
screen "3161_ParetoAlarmData" 1280x715, template "3xxx_Alarms&Events"
   Rectangle "recBaseScreenLocked" at 0,0 size 1280x708
      Visibility <- "bo_System_BaseScreenLocked"
   TextField "Text_SortBy" at 33,29 size 102x31; Text 'Sort By:'
   SymbolicIOField "List_ParetoSort" at 135,28 size 244x33; TextOn '1'; TextOff '0'; TextList "Pareto_Sort"
      ProcessValue <- "ParetoData_Sort"
   TextField "Title_Alarm" at 1,84 size 50x21; Text 'Alarm'
   TextField "Title_ID" at 63,84 size 24x21; Text 'ID'
   TextField "Title_Message" at 286,84 size 71x21; Text 'Meldung / Message'
   TextField "Title_TimesOccurred" at 516,67 size 76x38; Text 'Anzahl Time Occurred'
   TextField "Title_TotalDowntime" at 584,67 size 102x38; Text 'Unproduktiv Total Downtime'
   TextField "Title_MTTR" at 682,84 size 49x21; Text 'MTTR'
   TextField "Title_%" at 761,84 size 23x21; Text '%'
   TextField "Text_TotalUptime" at 842,192 size 119x40; Text 'Produktiv: [min] Total Uptime: [min]'
   TextField "Text_TotalDowntime" at 818,250 size 143x40; Text 'Unproduktiv: [min] Total Downtime: [min]'
   TextField "Text_PercentUptime" at 821,316 size 140x22; Text 'Produktiv in %: / Percent Uptime:'
   TextField "Text_TotalStops" at 855,374 size 106x22; Text 'Stopps: / Total Stops:'
   TextField "Text_MTTR" at 903,422 size 58x40; Text 'MTTR: [min]'
   TextField "Text_MTBF" at 904,480 size 57x40; Text 'MTBF: [min]'
   Button "Reset_Button" at 833,539 size 254x32; TextOff 'RESET'
      on Press: function_b14e0dd5("ParetoData_Reset", 0)
   IOField "TotalUptime" at 967,197 size 120x30; FormatPattern 9999.99
      ProcessValue <- "ParetoData_totalUptime"
   IOField "TotalDowntime" at 967,255 size 120x30; FormatPattern 9999.99
      ProcessValue <- "ParetoData_totalDowntime"
   IOField "PercentUptime" at 967,312 size 120x30; FormatPattern 999.9
      ProcessValue <- "ParetoData_percentUptime"
   IOField "TotalStops" at 967,370 size 120x30; FormatPattern 999
      ProcessValue <- "ParetoData_totalStops"
   IOField "MTTR" at 967,427 size 120x30; FormatPattern 9999.99
      ProcessValue <- "ParetoData_MTTR"
   IOField "MTBF" at 967,485 size 120x30; FormatPattern 9999.99
      ProcessValue <- "ParetoData_MTBF"
   TextField "Title_Alarm_1" at 14,118 size 29x31; Text '1:'
   TextField "Title_Alarm_2" at 14,166 size 29x31; Text '2:'
   TextField "Title_Alarm_3" at 14,214 size 29x31; Text '3:'
   TextField "Title_Alarm_4" at 14,262 size 29x31; Text '4:'
   TextField "Title_Alarm_5" at 14,310 size 29x31; Text '5:'
   TextField "Title_Alarm_6" at 14,358 size 29x31; Text '6:'
   TextField "Title_Alarm_7" at 14,406 size 29x31; Text '7:'
   TextField "Title_Alarm_8" at 14,454 size 29x31; Text '8:'
   TextField "Title_Alarm_9" at 14,502 size 29x31; Text '9:'
   TextField "Title_Alarm_10" at 6,550 size 44x31; Text '10:'
   TextField "Text_TotalTimeSinceReset" at 850,126 size 111x58; Text 'Zeit seit Rücksetzen: [min] Total Time Since Reset: [min]'
   IOField "TotalTimeSinceReset" at 967,140 size 120x30; FormatPattern 9999.99
      ProcessValue <- "ParetoData_totalTimeSinceReset"
   ScreenModuleView "ParetoFacePlate_1" at 49,115 size 760x38; ScreenModuleType ""
      Guid_{11997190-103935} <- "ParetoData_alarmOccurrence[1]"
   ScreenModuleView "ParetoFacePlate_2" at 49,163 size 760x38; ScreenModuleType ""
      Guid_{11997190-103935} <- "ParetoData_alarmOccurrence[2]"
   ScreenModuleView "ParetoFacePlate_3" at 49,211 size 760x38; ScreenModuleType ""
      Guid_{11997190-103935} <- "ParetoData_alarmOccurrence[3]"
   ScreenModuleView "ParetoFacePlate_4" at 49,259 size 760x38; ScreenModuleType ""
      Guid_{11997190-103935} <- "ParetoData_alarmOccurrence[4]"
   ScreenModuleView "ParetoFacePlate_5" at 49,307 size 760x38; ScreenModuleType ""
      Guid_{11997190-103935} <- "ParetoData_alarmOccurrence[5]"
   ScreenModuleView "ParetoFacePlate_6" at 49,355 size 760x38; ScreenModuleType ""
      Guid_{11997190-103935} <- "ParetoData_alarmOccurrence[6]"
   ScreenModuleView "ParetoFacePlate_7" at 49,403 size 760x38; ScreenModuleType ""
      Guid_{11997190-103935} <- "ParetoData_alarmOccurrence[7]"
   ScreenModuleView "ParetoFacePlate_8" at 49,451 size 760x38; ScreenModuleType ""
      Guid_{11997190-103935} <- "ParetoData_alarmOccurrence[8]"
   ScreenModuleView "ParetoFacePlate_9" at 49,499 size 760x38; ScreenModuleType ""
      Guid_{11997190-103935} <- "ParetoData_alarmOccurrence[9]"
   ScreenModuleView "ParetoFacePlate_10" at 49,547 size 760x38; ScreenModuleType ""
      Guid_{11997190-103935} <- "ParetoData_alarmOccurrence[10]"

screen "7001_RecipeControl" 1280x715, template "7xxx_Formats"
   Button "btn_Save" at 937,17 size 156x71; TextOff 'Save Current Recipe Datensatz Speichern Salvar'
      on Release: ResetBit("CPG_Recipe_Management.HMI_Command.Save.saveCmd")
      on Press: SetBit("CPG_Recipe_Management.HMI_Command.Save.saveCmd")
   Button "btn_Save_1" at 25,29 size 111x48; TextOff 'Reset All Times Rücksetzen Salvar'
      on Release: ResetBit("CPG_Recipe_Management.HMI_Command.resetAllTimes")
      on Press: SetBit("CPG_Recipe_Management.HMI_Command.resetAllTimes")
   Button "btn_Delete" at 444,538 size 150x45; TextOff 'Change Recipe Datensatz Ändern'
      on Release: ResetBit("CPG_Recipe_Management.HMI_Command.Change.changeCmd")
      on Press: SetBit("CPG_Recipe_Management.HMI_Command.Change.changeCmd")
   Button "btn_Rename" at 607,538 size 150x45; TextOff 'Save Recipe As Datensatz Speichern unter Rebautizar:'
      on Release: ResetBit("CPG_Recipe_Management.HMI_Command.Save.saveAsCmd")
      on Press: SetBit("CPG_Recipe_Management.HMI_Command.Save.saveAsCmd")
   Button "btn_WriteToPLC" at 771,538 size 150x45; TextOff 'Copy Recipe Datensatz Kopieren Write to PLC'
      on Release: ResetBit("CPG_Recipe_Management.HMI_Command.Copy.copyCmd")
      on Press: SetBit("CPG_Recipe_Management.HMI_Command.Copy.copyCmd")
   Button "btn_ReadFromPLC" at 935,538 size 150x45; TextOff 'Delete Recipe Datensatz Löschen Leer desde PLC'
      on Release: ResetBit("CPG_Recipe_Management.HMI_Command.Delete.deleteCmd")
      on Press: SetBit("CPG_Recipe_Management.HMI_Command.Delete.deleteCmd")
   Button "rec_BaseScreenLocked" at 0,0 size 1280x715; TextOff 'Text'
      Visibility <- "bo_System_BaseScreenLocked"
   IOField "I/O field_2" at 345,38 size 38x29; FormatPattern 999
      ProcessValue <- "CurrentRecipeID"
   TextField "Text field_5" at 166,39 size 157x27; Text 'Current Recipe: / Aktueller Datensatz:'
   IOField "I/O field_19" at 171,91 size 189x29; FormatPattern ????????????????????
      ProcessValue <- "CurrentRecipeName"
   TextField "Text field_26" at 8,84 size 156x48; Text 'Tap to Rename Current Recipe: Aktuellen Datensatz Umbenennen:'
   Button "Button_3" at 13,559 size 78x45; TextOff 'Text'; PictureOff "Up_Arrow"
      on Release: function_b9b71300("CPG_Recipe_Management.currentPages[4]", 1)
   Button "Button_4" at 117,559 size 78x45; TextOff 'Text'; PictureOff "Down_Arrow"
      on Release: function_dd21b452("CPG_Recipe_Management.currentPages[4]", 1)
   IOField "I/O field_30" at 293,571 size 35x21; FormatPattern 999
      ProcessValue <- "CPG_Recipe_Management.currentPages[4]"
   TextField "Text field_46" at 225,569 size 60x25; Text 'Page # / Seite #'
   TextField "Text field_47" at 337,569 size 32x25; Text 'of / von'
   IOField "I/O field_45" at 385,572 size 27x19; FormatPattern 999
      ProcessValue <- "CPG_Recipe_Management.maxPages[4]"
   Rectangle "Rectangle_7" at 438,24 size 224x56
      Visibility <- "RecipeChangeDisabled"
   TextField "Text field_45" at 455,28 size 190x48; Text 'Recipe changes disabled due to machine state Änderungen gesperrt wegen Maschinenzustand'
      Visibility <- "RecipeChangeDisabled"
   Rectangle "Rectangle_2" at 668,24 size 261x56
      Visibility <- "RecipeSetpointDiff"
   TextField "Text field_27" at 674,28 size 249x48; Text 'Warning: At least one value differs from the saved setpoints! Mindestens ein Wert entspricht nicht den Speicherwerten!'
      Visibility <- "RecipeSetpointDiff"
   Group "Group" at 5,531 size 421x27
   Group "Group_1" at 5,509 size 421x27
   Group "Group_3" at 5,488 size 421x27
   Group "Group_4" at 5,467 size 421x27
   Group "Group_6" at 5,446 size 421x27
   Group "Group_7" at 5,425 size 421x27
   Group "Group_8" at 5,404 size 421x27
   Group "Group_9" at 5,382 size 421x27
   Group "Group_10" at 5,361 size 421x27
   Group "Group_11" at 5,340 size 421x27
   Group "Group_12" at 5,319 size 421x27
   Group "Group_13" at 5,298 size 421x27
   Group "Group_14" at 5,277 size 421x27
   Group "Group_15" at 5,255 size 421x27
   Group "Group_16" at 5,234 size 421x27
   Group "Group_17" at 5,213 size 421x27
   Group "Group_18" at 5,192 size 421x27
   Group "Group_19" at 5,171 size 421x27
   Group "Group_20" at 5,150 size 421x27
   Group "Group_21" at 5,129 size 421x27
   IOField "I/O field_44" at 230,531 size 196x27; FormatPattern 9999999999999999999999999999999999999999
      ProcessValue <- "[19]"
      Visibility <- "[19]"
   IOField "I/O field_29" at 45,534 size 185x22; FormatPattern ????????????????????
      ProcessValue <- "[19]"
      Visibility <- "[19]"
   TextField "Text field_37" at 36,531 size 41x27; Text ':'
      Visibility <- "[19]"
   IOField "I/O field_65" at 5,531 size 37x27; FormatPattern 999
      ProcessValue <- "[19]"
      Visibility <- "[19]"
   IOField "I/O field_28" at 45,511 size 185x22; FormatPattern ????????????????????
      ProcessValue <- "[18]"
      Visibility <- "[18]"
   IOField "I/O field_43" at 230,509 size 196x27; FormatPattern 9999999999999999999999999999999999999999
      ProcessValue <- "[18]"
      Visibility <- "[18]"
   IOField "I/O field_64" at 5,509 size 37x27; FormatPattern 999
      ProcessValue <- "[18]"
      Visibility <- "[18]"
   TextField "Text field_36" at 36,509 size 41x27; Text ':'
      Visibility <- "[18]"
   IOField "I/O field_27" at 45,490 size 185x22; FormatPattern ????????????????????
      ProcessValue <- "[17]"
      Visibility <- "[17]"
   IOField "I/O field_42" at 230,488 size 196x27; FormatPattern 9999999999999999999999999999999999999999
      ProcessValue <- "[17]"
      Visibility <- "[17]"
   IOField "I/O field_63" at 5,488 size 37x27; FormatPattern 999
      ProcessValue <- "[17]"
      Visibility <- "[17]"
   TextField "Text field_35" at 36,488 size 41x27; Text ':'
      Visibility <- "[17]"
   IOField "I/O field_26" at 45,469 size 185x22; FormatPattern ????????????????????
      ProcessValue <- "[16]"
      Visibility <- "[16]"
   IOField "I/O field_41" at 230,467 size 196x27; FormatPattern 9999999999999999999999999999999999999999
      ProcessValue <- "[16]"
      Visibility <- "[16]"
   IOField "I/O field_62" at 5,467 size 37x27; FormatPattern 999
      ProcessValue <- "[16]"
      Visibility <- "[16]"
   TextField "Text field_34" at 36,467 size 41x27; Text ':'
      Visibility <- "[16]"
   IOField "I/O field_25" at 45,448 size 185x22; FormatPattern ????????????????????
      ProcessValue <- "[15]"
      Visibility <- "[15]"
   IOField "I/O field_40" at 230,446 size 196x27; FormatPattern 9999999999999999999999999999999999999999
      ProcessValue <- "[15]"
      Visibility <- "[15]"
   IOField "I/O field_61" at 5,446 size 37x27; FormatPattern 999
      ProcessValue <- "[15]"
      Visibility <- "[15]"
   TextField "Text field_33" at 36,446 size 41x27; Text ':'
      Visibility <- "[15]"
   IOField "I/O field_24" at 45,427 size 185x22; FormatPattern ????????????????????
      ProcessValue <- "[14]"
      Visibility <- "[14]"
   IOField "I/O field_39" at 230,425 size 196x27; FormatPattern 9999999999999999999999999999999999999999
      ProcessValue <- "[14]"
      Visibility <- "[14]"
   IOField "I/O field_60" at 5,425 size 37x27; FormatPattern 999
      ProcessValue <- "[14]"
      Visibility <- "[14]"
   TextField "Text field_32" at 36,425 size 41x27; Text ':'
      Visibility <- "[14]"
   IOField "I/O field_23" at 45,406 size 185x22; FormatPattern ????????????????????
      ProcessValue <- "[13]"
      Visibility <- "[13]"
   IOField "I/O field_38" at 230,404 size 196x27; FormatPattern 9999999999999999999999999999999999999999
      ProcessValue <- "[13]"
      Visibility <- "[13]"
   IOField "I/O field_59" at 5,404 size 37x27; FormatPattern 999
      ProcessValue <- "[13]"
      Visibility <- "[13]"
   TextField "Text field_31" at 36,404 size 41x27; Text ':'
      Visibility <- "[13]"
   IOField "I/O field_22" at 45,384 size 185x22; FormatPattern ????????????????????
      ProcessValue <- "[12]"
      Visibility <- "[12]"
   IOField "I/O field_32" at 230,382 size 196x27; FormatPattern 9999999999999999999999999999999999999999
      ProcessValue <- "[12]"
      Visibility <- "[12]"
   IOField "I/O field_58" at 5,382 size 37x27; FormatPattern 999
      ProcessValue <- "[12]"
      Visibility <- "[12]"
   TextField "Text field_30" at 36,382 size 41x27; Text ':'
      Visibility <- "[12]"
   IOField "I/O field_21" at 45,363 size 185x22; FormatPattern ????????????????????
      ProcessValue <- "[11]"
      Visibility <- "[11]"
   IOField "I/O field_37" at 230,361 size 196x27; FormatPattern 9999999999999999999999999999999999999999
      ProcessValue <- "[11]"
      Visibility <- "[11]"
   IOField "I/O field_57" at 5,361 size 37x27; FormatPattern 999
      ProcessValue <- "[11]"
      Visibility <- "[11]"
   TextField "Text field_29" at 36,361 size 41x27; Text ':'
      Visibility <- "[11]"
   IOField "I/O field_20" at 45,342 size 185x22; FormatPattern ????????????????????
      ProcessValue <- "[10]"
      Visibility <- "[10]"
   IOField "I/O field_36" at 230,340 size 196x27; FormatPattern 9999999999999999999999999999999999999999
      ProcessValue <- "[10]"
      Visibility <- "[10]"
   IOField "I/O field_56" at 5,340 size 37x27; FormatPattern 999
      ProcessValue <- "[10]"
      Visibility <- "[10]"
   TextField "Text field_28" at 36,340 size 41x27; Text ':'
      Visibility <- "[10]"
   IOField "I/O field_18" at 45,321 size 185x22; FormatPattern ????????????????????
      ProcessValue <- "[9]"
      Visibility <- "[9]"
   IOField "I/O field_35" at 230,319 size 196x27; FormatPattern 9999999999999999999999999999999999999999
      ProcessValue <- "[9]"
      Visibility <- "[9]"
   IOField "I/O field_55" at 5,319 size 37x27; FormatPattern 999
      ProcessValue <- "[9]"
      Visibility <- "[9]"
   TextField "Text field_25" at 36,319 size 41x27; Text ':'
      Visibility <- "[9]"
   IOField "I/O field_17" at 45,300 size 185x22; FormatPattern ????????????????????
      ProcessValue <- "[8]"
      Visibility <- "[8]"
   IOField "I/O field_34" at 230,298 size 196x27; FormatPattern 9999999999999999999999999999999999999999
      ProcessValue <- "[8]"
      Visibility <- "[8]"
   IOField "I/O field_54" at 5,298 size 37x27; FormatPattern 999
      ProcessValue <- "[8]"
      Visibility <- "[8]"
   TextField "Text field_24" at 36,298 size 41x27; Text ':'
      Visibility <- "[8]"
   IOField "I/O field_16" at 45,279 size 185x22; FormatPattern ????????????????????
      ProcessValue <- "[7]"
      Visibility <- "[7]"
   IOField "I/O field_33" at 230,277 size 196x27; FormatPattern 9999999999999999999999999999999999999999
      ProcessValue <- "[7]"
      Visibility <- "[7]"
   IOField "I/O field_53" at 5,277 size 37x27; FormatPattern 999
      ProcessValue <- "[7]"
      Visibility <- "[7]"
   TextField "Text field_23" at 36,277 size 41x27; Text ':'
      Visibility <- "[7]"
   IOField "I/O field_15" at 45,257 size 185x22; FormatPattern ????????????????????
      ProcessValue <- "[6]"
      Visibility <- "[6]"
   IOField "I/O field_31" at 230,255 size 196x27; FormatPattern 9999999999999999999999999999999999999999
      ProcessValue <- "[6]"
      Visibility <- "[6]"
   IOField "I/O field_52" at 5,255 size 37x27; FormatPattern 999
      ProcessValue <- "[6]"
      Visibility <- "[6]"
   TextField "Text field_22" at 36,255 size 41x27; Text ':'
      Visibility <- "[6]"
   IOField "I/O field_14" at 45,236 size 185x22; FormatPattern ????????????????????
      ProcessValue <- "[5]"
      Visibility <- "[5]"
   IOField "I/O field_8" at 230,234 size 196x27; FormatPattern 9999999999999999999999999999999999999999
      ProcessValue <- "[5]"
      Visibility <- "[5]"
   IOField "I/O field_51" at 5,234 size 37x27; FormatPattern 999
      ProcessValue <- "[5]"
      Visibility <- "[5]"
   TextField "Text field_21" at 36,234 size 41x27; Text ':'
      Visibility <- "[5]"
   IOField "I/O field_13" at 45,215 size 185x22; FormatPattern ????????????????????
      ProcessValue <- "[4]"
      Visibility <- "[4]"
   IOField "I/O field_7" at 230,213 size 196x27; FormatPattern 9999999999999999999999999999999999999999
      ProcessValue <- "[4]"
      Visibility <- "[4]"
   IOField "I/O field_50" at 5,213 size 37x27; FormatPattern 999
      ProcessValue <- "[4]"
      Visibility <- "[4]"
   TextField "Text field_20" at 36,213 size 41x27; Text ':'
      Visibility <- "[4]"
   IOField "I/O field_12" at 45,194 size 185x22; FormatPattern ????????????????????
      ProcessValue <- "[3]"
      Visibility <- "[3]"
   IOField "I/O field_6" at 230,192 size 196x27; FormatPattern 9999999999999999999999999999999999999999
      ProcessValue <- "[3]"
      Visibility <- "[3]"
   IOField "I/O field_49" at 5,192 size 37x27; FormatPattern 999
      ProcessValue <- "[3]"
      Visibility <- "[3]"
   TextField "Text field_19" at 36,192 size 41x27; Text ':'
      Visibility <- "[3]"
   IOField "I/O field_11" at 45,173 size 185x22; FormatPattern ????????????????????
      ProcessValue <- "[2]"
      Visibility <- "[2]"
   IOField "I/O field_4" at 230,171 size 196x27; FormatPattern 9999999999999999999999999999999999999999
      ProcessValue <- "[2]"
      Visibility <- "[2]"
   IOField "I/O field_48" at 5,171 size 37x27; FormatPattern 999
      ProcessValue <- "[2]"
      Visibility <- "[2]"
   TextField "Text field_18" at 36,171 size 41x27; Text ':'
      Visibility <- "[2]"
   IOField "I/O field_10" at 45,152 size 185x22; FormatPattern ????????????????????
      ProcessValue <- "[1]"
      Visibility <- "[1]"
   IOField "I/O field_5" at 230,150 size 196x27; FormatPattern 9999999999999999999999999999999999999999
      ProcessValue <- "[1]"
      Visibility <- "[1]"
   IOField "I/O field_47" at 5,150 size 37x27; FormatPattern 999
      ProcessValue <- "[1]"
      Visibility <- "[1]"
   TextField "Text field_17" at 36,150 size 41x27; Text ':'
      Visibility <- "[1]"
   IOField "I/O field_9" at 45,131 size 185x22; FormatPattern ????????????????????
      ProcessValue <- "[0]"
      Visibility <- "[0]"
   IOField "I/O field_3" at 230,129 size 196x27; FormatPattern 9999999999999999999999999999999999999999
      ProcessValue <- "[0]"
      Visibility <- "[0]"
   IOField "I/O field_46" at 5,129 size 37x27; FormatPattern 999
      ProcessValue <- "[0]"
      Visibility <- "[0]"
   TextField "Text field_16" at 36,129 size 41x27; Text ':'
      Visibility <- "[0]"
   Group "Group_26" at 560,148 size 446x339; FormatPattern ??????????????????????????????
   TextField "Text field_12" at 560,148 size 446x88; Text '"Save As" takes all running values - even those not saved - and saves them to the "Destination" recipe. To save to the current recipe, use the "Save" button in the upper right. "Speichern unter" übernimmt alle aktiven Werte, auch die ungespeicherten, und speichert sie in den "Ziel" Datensatz. Drücken Sie "Speichern" oben rechts, um den aktuellen Datensatz zu speichern.'
      Visibility <- "CPG_Recipe_Management.HMI_Indicator.saveAsConfirm"
   Button "Save Cancel" at 571,421 size 128x66; TextOff 'Cancel / Abbrechen'
      on Release: ResetBit("CPG_Recipe_Management.HMI_Command.Save.cancel")
      on Press: SetBit("CPG_Recipe_Management.HMI_Command.Save.cancel")
      Visibility <- "CPG_Recipe_Management.HMI_Indicator.saveAsConfirm"
   IOField "Save Name" at 630,362 size 285x29; FormatPattern ????????????????????
      Visibility <- "CPG_Recipe_Management.HMI_Indicator.saveAsConfirm"
      ProcessValue <- "CPG_Recipe_Management.HMI_Command.Save.saveAsNewName"
   Button "Save Req" at 847,421 size 128x66; TextOff 'Continue Save As Fortsetzen Speichern unter'
      on Release: ResetBit("CPG_Recipe_Management.HMI_Command.Save.request")
      on Press: SetBit("CPG_Recipe_Management.HMI_Command.Save.request")
      Visibility <- "CPG_Recipe_Management.HMI_Indicator.saveAsConfirm"
   IOField "Save Destination" at 912,291 size 37x27; FormatPattern 999
      ProcessValue <- "CPG_Recipe_Management.HMI_Command.Save.saveAsDestinationID"
      Visibility <- "CPG_Recipe_Management.HMI_Indicator.saveAsConfirm"
   TextField "Text field_14" at 806,295 size 97x25; Text 'Destination: / Ziel:'
      Visibility <- "CPG_Recipe_Management.HMI_Indicator.saveAsConfirm"
   TextField "Text field_13" at 605,295 size 181x25; Text 'Source: Current Values / Quelle: Aktuelle Werte'
      Visibility <- "CPG_Recipe_Management.HMI_Indicator.saveAsConfirm"
   TextField "Text field_42" at 666,334 size 319x25; Text 'New name for saved recipe: / Neuer Name für gespeicherten Datensatz:'
      Visibility <- "CPG_Recipe_Management.HMI_Indicator.saveAsConfirm"
   Group "Group_25" at 847,421 size 128x66
   Rectangle "Rectangle_4" at 847,421 size 128x66
      Visibility <- "CPG_Recipe_Management.HMI_Indicator.saveAsErr"
   TextField "Text field_41" at 862,431 size 106x46; Text 'Cannot Save Invalid ID Nicht möglich Ungültige ID'
      Visibility <- "CPG_Recipe_Management.HMI_Indicator.saveAsErr"
   Group "Group_5" at 571,159 size 404x328; FormatPattern 99
   Button "Button_1" at 571,421 size 128x66; TextOff 'Cancel / Abbrechen'
      on Release: ResetBit("CPG_Recipe_Management.HMI_Command.Change.cancel")
      on Press: SetBit("CPG_Recipe_Management.HMI_Command.Change.cancel")
      Visibility <- "CPG_Recipe_Management.HMI_Indicator.changeConfirm"
   Button "Button_2" at 847,421 size 128x66; TextOff 'Continue Change Fortsetzen Ändern'
      on Release: ResetBit("CPG_Recipe_Management.HMI_Command.Change.request")
      on Press: SetBit("CPG_Recipe_Management.HMI_Command.Change.request")
      Visibility <- "CPG_Recipe_Management.HMI_Indicator.changeConfirm"
   TextField "Text field_4" at 581,352 size 376x46; Text 'Are you sure you want to change recipes and lose any unsaved data? Wollen Sie den Datensatz ändern? Ungespeicherte Daten gehen verloren.'
      Visibility <- "CPG_Recipe_Management.HMI_Indicator.changeConfirm"
   IOField "I/O field_1" at 676,291 size 37x27; FormatPattern 999
      Visibility <- "CPG_Recipe_Management.HMI_Indicator.changeConfirm"
      ProcessValue <- "CPG_Recipe_Management.HMI_Command.Change.changeID"
   TextField "Text field_2" at 605,295 size 62x25; Text 'Source: / Quelle:'
      Visibility <- "CPG_Recipe_Management.HMI_Indicator.changeConfirm"
   TextField "Text field_3" at 725,295 size 216x25; Text 'Destination: Current Values / Ziel: Aktuelle Werte'
      Visibility <- "CPG_Recipe_Management.HMI_Indicator.changeConfirm"
   TextField "Text field_1" at 604,159 size 327x88; Text '"Change" (Load) sets the current values equal to the values saved in "Source". Any unsaved data is lost. "Ändern" (Laden) setzt die aktuellen Werte gleich den Werten in "Quelle". Nicht gespeicherte Daten gehen verloren.'
      Visibility <- "CPG_Recipe_Management.HMI_Indicator.changeConfirm"
   Rectangle "Rectangle_6" at 847,421 size 128x66
      Visibility <- "CPG_Recipe_Management.HMI_Indicator.changeErr"
   TextField "Text field_44" at 852,431 size 118x46; Text 'Cannot Change Invalid ID Nicht möglich Ungültige ID'
      Visibility <- "CPG_Recipe_Management.HMI_Indicator.changeErr"
   Group "Group_22" at 560,148 size 428x339; FormatPattern ??????????????????????????????
   Button "Copy Req" at 847,421 size 128x66; TextOff 'Continue Copy Fortsetzen Kopieren'
      on Release: ResetBit("CPG_Recipe_Management.HMI_Command.Copy.request")
      on Press: SetBit("CPG_Recipe_Management.HMI_Command.Copy.request")
      Visibility <- "CPG_Recipe_Management.HMI_Indicator.copyConfirm"
   IOField "Copy Name" at 630,362 size 285x29; FormatPattern ????????????????????
      ProcessValue <- "CPG_Recipe_Management.HMI_Command.Copy.copyNewName"
      Visibility <- "CPG_Recipe_Management.HMI_Indicator.copyConfirm"
   TextField "Text field_15" at 685,334 size 194x25; Text 'Recipe Name for Copy: / Datensatz zum Kopieren:'
      Visibility <- "CPG_Recipe_Management.HMI_Indicator.copyConfirm"
   TextField "Text field_8" at 560,148 size 428x88; Text '"Copy" all of the saved values in "Source" to a different recipe at "Destination". Using this option only copies the saved values. The "Destination" must not be the current recipe. "Kopieren" aller gespeicherten Werte in "Quelle" in einen anderen Datensatz unter "Ziel". Mit dieser Option werden nur die gespeicherten Werte kopiert. Das "Ziel" darf nicht der aktuelle Datensatz sein.'
      Visibility <- "CPG_Recipe_Management.HMI_Indicator.copyConfirm"
   Button "Copy Cancel" at 571,421 size 128x66; TextOff 'Cancel / Abbrechen'
      on Release: ResetBit("CPG_Recipe_Management.HMI_Command.Copy.cancel")
      on Press: SetBit("CPG_Recipe_Management.HMI_Command.Copy.cancel")
      Visibility <- "CPG_Recipe_Management.HMI_Indicator.copyConfirm"
   TextField "Text field_10" at 605,295 size 62x25; Text 'Source: / Quelle:'
      Visibility <- "CPG_Recipe_Management.HMI_Indicator.copyConfirm"
   IOField "Copy Source" at 676,291 size 37x27; FormatPattern 999
      ProcessValue <- "CPG_Recipe_Management.HMI_Command.Copy.copySourceID"
      Visibility <- "CPG_Recipe_Management.HMI_Indicator.copyConfirm"
   TextField "Text field_11" at 806,295 size 97x25; Text 'Destination: / Ziel:'
      Visibility <- "CPG_Recipe_Management.HMI_Indicator.copyConfirm"
   IOField "Copy Destination" at 912,291 size 37x27; FormatPattern 999
      ProcessValue <- "CPG_Recipe_Management.HMI_Command.Copy.copyDestinationID"
      Visibility <- "CPG_Recipe_Management.HMI_Indicator.copyConfirm"
   Group "Group_2" at 847,421 size 128x66
   Rectangle "Rectangle_3" at 847,421 size 128x66
      Visibility <- "CPG_Recipe_Management.HMI_Indicator.copyErr"
   TextField "Text field_39" at 862,431 size 107x46; Text 'Cannot Copy Invalid IDs Nicht möglich Ungültige IDs'
      Visibility <- "CPG_Recipe_Management.HMI_Indicator.copyErr"
   Group "Group_24" at 554,155 size 529x332; FormatPattern 99
   TextField "Text field_6" at 554,155 size 529x67; Text '"Delete" sets the values of a saved recipe to their defaults, usually zero or null. It also deletes the recipe name. You cannot delete the currently loaded recipe. "Löschen" initialisiert die Werte eines vorhandenen Datensatzes, üblicherweise 0 oder Leer. Es wird auch der Datensatzname gelöscht. Der aktive Datensatz kann nicht gelöscht werden.'
      Visibility <- "CPG_Recipe_Management.HMI_Indicator.deleteConfirm"
   TextField "Text field_9" at 610,347 size 357x46; Text 'Are you sure you want to delete this recipe and lose any unsaved data? Sind Sie sicher dass Sie das Löschen abbrechen wollen? Ungespeicherte Daten gehen verloren.'
      Visibility <- "CPG_Recipe_Management.HMI_Indicator.deleteConfirm"
   Button "Delete Cancel" at 571,421 size 128x66; TextOff 'Cancel / Abbrechen'
      on Release: ResetBit("CPG_Recipe_Management.HMI_Command.Delete.cancel")
      on Press: SetBit("CPG_Recipe_Management.HMI_Command.Delete.cancel")
      Visibility <- "CPG_Recipe_Management.HMI_Indicator.deleteConfirm"
   Button "Delete Req" at 847,421 size 128x66; TextOff 'Continue Delete Fortsetzen Löschen'
      on Release: ResetBit("CPG_Recipe_Management.HMI_Command.Delete.request")
      on Press: SetBit("CPG_Recipe_Management.HMI_Command.Delete.request")
      Visibility <- "CPG_Recipe_Management.HMI_Indicator.deleteConfirm"
   TextField "Text field_7" at 686,295 size 136x25; Text 'Recipe to Delete: / Datensatz:'
      Visibility <- "CPG_Recipe_Management.HMI_Indicator.deleteConfirm"
   IOField "Delete Destination" at 831,291 size 37x27; FormatPattern 999
      ProcessValue <- "CPG_Recipe_Management.HMI_Command.Delete.deleteID"
      Visibility <- "CPG_Recipe_Management.HMI_Indicator.deleteConfirm"
   Group "Group_23" at 847,421 size 128x66
   Rectangle "Rectangle_5" at 847,421 size 128x66
      Visibility <- "CPG_Recipe_Management.HMI_Indicator.deleteErr"
   TextField "Text field_43" at 855,431 size 112x46; Text 'Cannot Delete Invalid ID Nicht möglich Ungültige ID'
      Visibility <- "CPG_Recipe_Management.HMI_Indicator.deleteErr"

screen "7041_RecipeSetpoints_REAL" 1280x715, template "7xxx_Formats"
   Button "rec_BaseScreenLocked" at 0,0 size 1280x715; TextOff 'Text'
      Visibility <- "bo_System_BaseScreenLocked"
   ScreenModuleView "Setpoint_Display_Real_2" at 4,166 size 1090x44; ScreenModuleType ""
      on Guid_{11997190-50501}: function_efd93a16("pop_recipes_REAL", 200, 50, -1, -1, 1); SetTag("CPG_Recipe_Management.popupTrackers[0]", 1)
      Guid_{11997190-47977} <- "CPG_Recipe_Management.setpointsArray_REAL[1]"
      Guid_{11997190-73128} <- "[1]"
   ScreenModuleView "Setpoint_Display_Real_1" at 4,132 size 1090x44; ScreenModuleType ""
      on Guid_{11997190-50501}: function_efd93a16("pop_recipes_REAL", 200, 50, -1, -1, 1); SetTag("CPG_Recipe_Management.popupTrackers[0]", 0)
      Guid_{11997190-47977} <- "CPG_Recipe_Management.setpointsArray_REAL[0]"
      Guid_{11997190-73128} <- "[0]"
   ScreenModuleView "Setpoint_Display_Real_3" at 4,200 size 1090x44; ScreenModuleType ""
      on Guid_{11997190-50501}: function_efd93a16("pop_recipes_REAL", 200, 50, -1, -1, 1); SetTag("CPG_Recipe_Management.popupTrackers[0]", 2)
      Guid_{11997190-47977} <- "CPG_Recipe_Management.setpointsArray_REAL[2]"
      Guid_{11997190-73128} <- "[2]"
   ScreenModuleView "Setpoint_Display_Real_4" at 4,234 size 1090x44; ScreenModuleType ""
      on Guid_{11997190-50501}: function_efd93a16("pop_recipes_REAL", 200, 50, -1, -1, 1); SetTag("CPG_Recipe_Management.popupTrackers[0]", 3)
      Guid_{11997190-47977} <- "CPG_Recipe_Management.setpointsArray_REAL[3]"
      Guid_{11997190-73128} <- "[3]"
   ScreenModuleView "Setpoint_Display_Real_5" at 4,268 size 1090x44; ScreenModuleType ""
      on Guid_{11997190-50501}: function_efd93a16("pop_recipes_REAL", 200, 50, -1, -1, 1); SetTag("CPG_Recipe_Management.popupTrackers[0]", 4)
      Guid_{11997190-47977} <- "CPG_Recipe_Management.setpointsArray_REAL[4]"
      Guid_{11997190-73128} <- "[4]"
   ScreenModuleView "Setpoint_Display_Real_6" at 4,302 size 1090x44; ScreenModuleType ""
      on Guid_{11997190-50501}: function_efd93a16("pop_recipes_REAL", 200, 50, -1, -1, 1); SetTag("CPG_Recipe_Management.popupTrackers[0]", 5)
      Guid_{11997190-47977} <- "CPG_Recipe_Management.setpointsArray_REAL[5]"
      Guid_{11997190-73128} <- "[5]"
   ScreenModuleView "Setpoint_Display_Real_7" at 4,336 size 1090x44; ScreenModuleType ""
      on Guid_{11997190-50501}: function_efd93a16("pop_recipes_REAL", 200, 50, -1, -1, 1); SetTag("CPG_Recipe_Management.popupTrackers[0]", 6)
      Guid_{11997190-47977} <- "CPG_Recipe_Management.setpointsArray_REAL[6]"
      Guid_{11997190-73128} <- "[6]"
   ScreenModuleView "Setpoint_Display_Real_8" at 4,370 size 1090x44; ScreenModuleType ""
      on Guid_{11997190-50501}: function_efd93a16("pop_recipes_REAL", 200, 50, -1, -1, 1); SetTag("CPG_Recipe_Management.popupTrackers[0]", 7)
      Guid_{11997190-47977} <- "CPG_Recipe_Management.setpointsArray_REAL[7]"
      Guid_{11997190-73128} <- "[7]"
   ScreenModuleView "Setpoint_Display_Real_9" at 4,404 size 1090x44; ScreenModuleType ""
      on Guid_{11997190-50501}: function_efd93a16("pop_recipes_REAL", 200, 50, -1, -1, 1); SetTag("CPG_Recipe_Management.popupTrackers[0]", 8)
      Guid_{11997190-47977} <- "CPG_Recipe_Management.setpointsArray_REAL[8]"
      Guid_{11997190-73128} <- "[8]"
   ScreenModuleView "Setpoint_Display_Real_10" at 4,438 size 1090x44; ScreenModuleType ""
      on Guid_{11997190-50501}: function_efd93a16("pop_recipes_REAL", 200, 50, -1, -1, 1); SetTag("CPG_Recipe_Management.popupTrackers[0]", 9)
      Guid_{11997190-47977} <- "CPG_Recipe_Management.setpointsArray_REAL[9]"
      Guid_{11997190-73128} <- "[9]"
   ScreenModuleView "Setpoint_Display_Real_11" at 4,472 size 1090x44; ScreenModuleType ""
      on Guid_{11997190-50501}: function_efd93a16("pop_recipes_REAL", 200, 50, -1, -1, 1); SetTag("CPG_Recipe_Management.popupTrackers[0]", 10)
      Guid_{11997190-47977} <- "CPG_Recipe_Management.setpointsArray_REAL[10]"
      Guid_{11997190-73128} <- "[10]"
   ScreenModuleView "Setpoint_Display_Real_12" at 4,506 size 1090x44; ScreenModuleType ""
      on Guid_{11997190-50501}: function_efd93a16("pop_recipes_REAL", 200, 50, -1, -1, 1); SetTag("CPG_Recipe_Management.popupTrackers[0]", 11)
      Guid_{11997190-47977} <- "CPG_Recipe_Management.setpointsArray_REAL[11]"
      Guid_{11997190-73128} <- "[11]"
   TextField "Text field_2" at 35,93 size 115x25; Text 'Setpoint Name / Sollwert-Name'
   TextField "Text field_6" at 243,83 size 72x46; Text 'Current Value Aktueller Wert'
   TextField "Text field_7" at 384,93 size 32x25; Text 'Min'
   TextField "Text field_4" at 506,93 size 36x25; Text 'Max'
   IOField "I/O field_9" at 757,42 size 53x36; FormatPattern 999
      ProcessValue <- "RecipeID_A"
   IOField "I/O field_10" at 883,42 size 53x36; FormatPattern 999
      ProcessValue <- "RecipeID_B"
   IOField "I/O field_11" at 998,42 size 53x36; FormatPattern 999
      ProcessValue <- "RecipeID_C"
   IOField "I/O field_13" at 550,83 size 187x22; FormatPattern ????????????????????
      ProcessValue <- "CurrentRecipeName"
   IOField "I/O field_14" at 907,104 size 187x22; FormatPattern ????????????????????
      ProcessValue <- "RecipeName_C"
   IOField "I/O field_15" at 816,83 size 187x22; FormatPattern ????????????????????
      ProcessValue <- "RecipeName_B"
   IOField "I/O field_16" at 690,103 size 187x23; FormatPattern ????????????????????
      ProcessValue <- "RecipeName_A"
   TextField "Text field_1" at 748,15 size 98x25; Text 'Recipe A / Datensatz A'
   TextField "Text field_3" at 874,15 size 97x25; Text 'Recipe B / Datensatz B'
   TextField "Text field_8" at 989,15 size 97x25; Text 'Recipe C / Datensatz C'
   TextField "Text field_9" at 125,40 size 209x25; Text 'RECIPE SETPOINTS - REAL / Rezeptur Sollwerte - REAL'
   Button "Button_1" at 160,555 size 78x45; TextOff 'Text'; PictureOff "Up_Arrow"
      on Release: function_b9b71300("CPG_Recipe_Management.currentPages[0]", 1)
   Button "Button_2" at 287,555 size 78x45; TextOff 'Text'; PictureOff "Down_Arrow"
      on Release: function_dd21b452("CPG_Recipe_Management.currentPages[0]", 1)
   TextField "Text field_10" at 35,565 size 126x25; Text 'Pg Up/Down / Seite vor/zurück'
   IOField "I/O field_1" at 446,565 size 35x25; FormatPattern 999
      ProcessValue <- "CPG_Recipe_Management.currentPages[0]"
   TextField "Text field_11" at 381,565 size 60x25; Text 'Page # / Seite #'
   TextField "Text field_12" at 488,565 size 32x25; Text 'of / von'
   IOField "I/O field_2" at 534,564 size 37x27; FormatPattern 999
      ProcessValue <- "CPG_Recipe_Management.maxPages[0]"
   Group "Group" at 588,37 size 110x46
   TextField "Text field_5" at 588,37 size 88x46; Text 'Current Recipe: Aktueller Datensatz:'
   IOField "I/O field_12" at 663,48 size 35x25; FormatPattern 999
      ProcessValue <- "CurrentRecipeID"

screen "7081_RecipeSetpoints_DINT" 1280x715, template "7xxx_Formats"
   Button "rec_BaseScreenLocked" at 0,0 size 1280x715; TextOff 'Text'
      Visibility <- "bo_System_BaseScreenLocked"
   ScreenModuleView "Setpoint_Display_Dint_3" at 4,200 size 1090x44; ScreenModuleType ""
      on Guid_{11997190-50501}: function_efd93a16("pop_recipes_DINT", 200, 50, -1, -1, 1); SetTag("CPG_Recipe_Management.popupTrackers[1]", 2)
      Guid_{11997190-47977} <- "CPG_Recipe_Management.setpointsArray_DINT[2]"
      Guid_{11997190-75846} <- "[2]"
   ScreenModuleView "Setpoint_Display_Dint_1" at 4,132 size 1090x44; ScreenModuleType ""
      on Guid_{11997190-50501}: function_efd93a16("pop_recipes_DINT", 200, 50, -1, -1, 1); SetTag("CPG_Recipe_Management.popupTrackers[1]", 0)
      Guid_{11997190-47977} <- "CPG_Recipe_Management.setpointsArray_DINT[0]"
      Guid_{11997190-75846} <- "[0]"
   ScreenModuleView "Setpoint_Display_Dint_2" at 4,166 size 1090x44; ScreenModuleType ""
      on Guid_{11997190-50501}: function_efd93a16("pop_recipes_DINT", 200, 50, -1, -1, 1); SetTag("CPG_Recipe_Management.popupTrackers[1]", 1)
      Guid_{11997190-47977} <- "CPG_Recipe_Management.setpointsArray_DINT[1]"
      Guid_{11997190-75846} <- "[1]"
   ScreenModuleView "Setpoint_Display_Dint_4" at 4,234 size 1090x44; ScreenModuleType ""
      on Guid_{11997190-50501}: function_efd93a16("pop_recipes_DINT", 200, 50, -1, -1, 1); SetTag("CPG_Recipe_Management.popupTrackers[1]", 3)
      Guid_{11997190-47977} <- "CPG_Recipe_Management.setpointsArray_DINT[3]"
      Guid_{11997190-75846} <- "[3]"
   ScreenModuleView "Setpoint_Display_Dint_5" at 4,268 size 1090x44; ScreenModuleType ""
      on Guid_{11997190-50501}: function_efd93a16("pop_recipes_DINT", 200, 50, -1, -1, 1); SetTag("CPG_Recipe_Management.popupTrackers[1]", 4)
      Guid_{11997190-47977} <- "CPG_Recipe_Management.setpointsArray_DINT[4]"
      Guid_{11997190-75846} <- "[4]"
   ScreenModuleView "Setpoint_Display_Dint_6" at 4,302 size 1090x44; ScreenModuleType ""
      on Guid_{11997190-50501}: function_efd93a16("pop_recipes_DINT", 200, 50, -1, -1, 1); SetTag("CPG_Recipe_Management.popupTrackers[1]", 5)
      Guid_{11997190-47977} <- "CPG_Recipe_Management.setpointsArray_DINT[5]"
      Guid_{11997190-75846} <- "[5]"
   ScreenModuleView "Setpoint_Display_Dint_7" at 4,336 size 1090x44; ScreenModuleType ""
      on Guid_{11997190-50501}: function_efd93a16("pop_recipes_DINT", 200, 50, -1, -1, 1); SetTag("CPG_Recipe_Management.popupTrackers[1]", 6)
      Guid_{11997190-47977} <- "CPG_Recipe_Management.setpointsArray_DINT[6]"
      Guid_{11997190-75846} <- "[6]"
   ScreenModuleView "Setpoint_Display_Dint_8" at 4,370 size 1090x44; ScreenModuleType ""
      on Guid_{11997190-50501}: function_efd93a16("pop_recipes_DINT", 200, 50, -1, -1, 1); SetTag("CPG_Recipe_Management.popupTrackers[1]", 7)
      Guid_{11997190-47977} <- "CPG_Recipe_Management.setpointsArray_DINT[7]"
      Guid_{11997190-75846} <- "[7]"
   ScreenModuleView "Setpoint_Display_Dint_9" at 4,404 size 1090x44; ScreenModuleType ""
      on Guid_{11997190-50501}: function_efd93a16("pop_recipes_DINT", 200, 50, -1, -1, 1); SetTag("CPG_Recipe_Management.popupTrackers[1]", 8)
      Guid_{11997190-47977} <- "CPG_Recipe_Management.setpointsArray_DINT[8]"
      Guid_{11997190-75846} <- "[8]"
   ScreenModuleView "Setpoint_Display_Dint_10" at 4,438 size 1090x44; ScreenModuleType ""
      on Guid_{11997190-50501}: function_efd93a16("pop_recipes_DINT", 200, 50, -1, -1, 1); SetTag("CPG_Recipe_Management.popupTrackers[1]", 9)
      Guid_{11997190-47977} <- "CPG_Recipe_Management.setpointsArray_DINT[9]"
      Guid_{11997190-75846} <- "[9]"
   ScreenModuleView "Setpoint_Display_Dint_11" at 4,472 size 1090x44; ScreenModuleType ""
      on Guid_{11997190-50501}: function_efd93a16("pop_recipes_DINT", 200, 50, -1, -1, 1); SetTag("CPG_Recipe_Management.popupTrackers[1]", 10)
      Guid_{11997190-47977} <- "CPG_Recipe_Management.setpointsArray_DINT[10]"
      Guid_{11997190-75846} <- "[10]"
   ScreenModuleView "Setpoint_Display_Dint_12" at 4,506 size 1090x44; ScreenModuleType ""
      on Guid_{11997190-50501}: function_efd93a16("pop_recipes_DINT", 200, 50, -1, -1, 1); SetTag("CPG_Recipe_Management.popupTrackers[1]", 11)
      Guid_{11997190-47977} <- "CPG_Recipe_Management.setpointsArray_DINT[11]"
      Guid_{11997190-75846} <- "[11]"
   TextField "Text field_9" at 125,40 size 208x25; Text 'RECIPE SETPOINTS - DINT / Rezeptur Sollwerte - DINT'
   Button "Button_3" at 160,555 size 78x45; TextOff 'Text'; PictureOff "Up_Arrow"
      on Release: function_b9b71300("CPG_Recipe_Management.currentPages[1]", 1)
   Button "Button_4" at 287,555 size 78x45; TextOff 'Text'; PictureOff "Down_Arrow"
      on Release: function_dd21b452("CPG_Recipe_Management.currentPages[1]", 1)
   TextField "Text field_10" at 35,565 size 126x25; Text 'Pg Up/Down / Seite vor/zurück'
   IOField "I/O field_3" at 446,565 size 35x25; FormatPattern 999
      ProcessValue <- "CPG_Recipe_Management.currentPages[1]"
   TextField "Text field_13" at 381,565 size 60x25; Text 'Page # / Seite #'
   TextField "Text field_14" at 488,565 size 32x25; Text 'of / von'
   IOField "I/O field_4" at 534,564 size 37x27; FormatPattern 999
      ProcessValue <- "CPG_Recipe_Management.maxPages[1]"
   TextField "Text field_2" at 35,93 size 115x25; Text 'Setpoint Name / Sollwert-Name'
   TextField "Text field_6" at 243,83 size 72x46; Text 'Current Value Aktueller Wert'
   TextField "Text field_7" at 384,93 size 32x25; Text 'Min'
   TextField "Text field_4" at 506,93 size 36x25; Text 'Max'
   IOField "I/O field_9" at 757,42 size 53x36; FormatPattern 999
      ProcessValue <- "RecipeID_A"
   IOField "I/O field_10" at 883,42 size 53x36; FormatPattern 999
      ProcessValue <- "RecipeID_B"
   IOField "I/O field_11" at 998,42 size 53x36; FormatPattern 999
      ProcessValue <- "RecipeID_C"
   IOField "I/O field_13" at 550,83 size 187x22; FormatPattern ????????????????????
      ProcessValue <- "CurrentRecipeName"
   IOField "I/O field_14" at 907,104 size 187x22; FormatPattern ????????????????????
      ProcessValue <- "RecipeName_C"
   IOField "I/O field_15" at 816,83 size 187x22; FormatPattern ????????????????????
      ProcessValue <- "RecipeName_B"
   IOField "I/O field_16" at 690,103 size 187x23; FormatPattern ????????????????????
      ProcessValue <- "RecipeName_A"
   TextField "Text field_1" at 748,15 size 98x25; Text 'Recipe A / Datensatz A'
   TextField "Text field_3" at 874,15 size 97x25; Text 'Recipe B / Datensatz B'
   TextField "Text field_8" at 989,15 size 97x25; Text 'Recipe C / Datensatz C'
   Group "Group" at 588,37 size 110x46
   TextField "Text field_5" at 588,37 size 88x46; Text 'Current Recipe: Aktueller Datensatz:'
   IOField "I/O field_12" at 663,48 size 35x25; FormatPattern 999
      ProcessValue <- "CurrentRecipeID"

screen "7121_RecipeSetpoints_BOOL" 1280x715, template "7xxx_Formats"
   Button "rec_BaseScreenLocked" at 0,0 size 1280x715; TextOff 'Text'
      Visibility <- "bo_System_BaseScreenLocked"
   ScreenModuleView "Setpoint_Display_3" at 4,200 size 1090x44; ScreenModuleType ""
      on Guid_{11997190-50501}: function_efd93a16("pop_recipes_BOOL", 200, 50, -1, -1, 1); SetTag("CPG_Recipe_Management.popupTrackers[2]", 2)
      Guid_{11997190-47977} <- "CPG_Recipe_Management.setpointsArray_BOOL[2]"
      Guid_{11997190-76108} <- "[2]"
   ScreenModuleView "Setpoint_Display_1" at 4,132 size 1090x44; ScreenModuleType ""
      on Guid_{11997190-50501}: function_efd93a16("pop_recipes_BOOL", 200, 50, -1, -1, 1); SetTag("CPG_Recipe_Management.popupTrackers[2]", 0)
      Guid_{11997190-47977} <- "CPG_Recipe_Management.setpointsArray_BOOL[0]"
      Guid_{11997190-76108} <- "[0]"
   ScreenModuleView "Setpoint_Display_2" at 4,166 size 1090x44; ScreenModuleType ""
      on Guid_{11997190-50501}: function_efd93a16("pop_recipes_BOOL", 200, 50, -1, -1, 1); SetTag("CPG_Recipe_Management.popupTrackers[2]", 1)
      Guid_{11997190-47977} <- "CPG_Recipe_Management.setpointsArray_BOOL[1]"
      Guid_{11997190-76108} <- "[1]"
   ScreenModuleView "Setpoint_Display_4" at 4,234 size 1090x44; ScreenModuleType ""
      on Guid_{11997190-50501}: function_efd93a16("pop_recipes_BOOL", 200, 50, -1, -1, 1); SetTag("CPG_Recipe_Management.popupTrackers[2]", 3)
      Guid_{11997190-47977} <- "CPG_Recipe_Management.setpointsArray_BOOL[3]"
      Guid_{11997190-76108} <- "[3]"
   ScreenModuleView "Setpoint_Display_5" at 4,268 size 1090x44; ScreenModuleType ""
      on Guid_{11997190-50501}: function_efd93a16("pop_recipes_BOOL", 200, 50, -1, -1, 1); SetTag("CPG_Recipe_Management.popupTrackers[2]", 4)
      Guid_{11997190-47977} <- "CPG_Recipe_Management.setpointsArray_BOOL[4]"
      Guid_{11997190-76108} <- "[4]"
   ScreenModuleView "Setpoint_Display_6" at 4,302 size 1090x44; ScreenModuleType ""
      on Guid_{11997190-50501}: function_efd93a16("pop_recipes_BOOL", 200, 50, -1, -1, 1); SetTag("CPG_Recipe_Management.popupTrackers[2]", 5)
      Guid_{11997190-47977} <- "CPG_Recipe_Management.setpointsArray_BOOL[5]"
      Guid_{11997190-76108} <- "[5]"
   ScreenModuleView "Setpoint_Display_7" at 4,336 size 1090x44; ScreenModuleType ""
      on Guid_{11997190-50501}: function_efd93a16("pop_recipes_BOOL", 200, 50, -1, -1, 1); SetTag("CPG_Recipe_Management.popupTrackers[2]", 6)
      Guid_{11997190-47977} <- "CPG_Recipe_Management.setpointsArray_BOOL[6]"
      Guid_{11997190-76108} <- "[6]"
   ScreenModuleView "Setpoint_Display_8" at 4,370 size 1090x44; ScreenModuleType ""
      on Guid_{11997190-50501}: function_efd93a16("pop_recipes_BOOL", 200, 50, -1, -1, 1); SetTag("CPG_Recipe_Management.popupTrackers[2]", 7)
      Guid_{11997190-47977} <- "CPG_Recipe_Management.setpointsArray_BOOL[7]"
      Guid_{11997190-76108} <- "[7]"
   ScreenModuleView "Setpoint_Display_9" at 4,404 size 1090x44; ScreenModuleType ""
      on Guid_{11997190-50501}: function_efd93a16("pop_recipes_BOOL", 200, 50, -1, -1, 1); SetTag("CPG_Recipe_Management.popupTrackers[2]", 8)
      Guid_{11997190-47977} <- "CPG_Recipe_Management.setpointsArray_BOOL[8]"
      Guid_{11997190-76108} <- "[8]"
   ScreenModuleView "Setpoint_Display_10" at 4,438 size 1090x44; ScreenModuleType ""
      on Guid_{11997190-50501}: function_efd93a16("pop_recipes_BOOL", 200, 50, -1, -1, 1); SetTag("CPG_Recipe_Management.popupTrackers[2]", 9)
      Guid_{11997190-47977} <- "CPG_Recipe_Management.setpointsArray_BOOL[9]"
      Guid_{11997190-76108} <- "[9]"
   ScreenModuleView "Setpoint_Display_11" at 4,472 size 1090x44; ScreenModuleType ""
      on Guid_{11997190-50501}: function_efd93a16("pop_recipes_BOOL", 200, 50, -1, -1, 1); SetTag("CPG_Recipe_Management.popupTrackers[2]", 10)
      Guid_{11997190-47977} <- "CPG_Recipe_Management.setpointsArray_BOOL[10]"
      Guid_{11997190-76108} <- "[10]"
   ScreenModuleView "Setpoint_Display_12" at 4,506 size 1090x44; ScreenModuleType ""
      on Guid_{11997190-50501}: function_efd93a16("pop_recipes_BOOL", 200, 50, -1, -1, 1); SetTag("CPG_Recipe_Management.popupTrackers[2]", 11)
      Guid_{11997190-47977} <- "CPG_Recipe_Management.setpointsArray_BOOL[11]"
      Guid_{11997190-76108} <- "[11]"
   TextField "Text field_9" at 125,40 size 211x25; Text 'RECIPE SETPOINTS - BOOL / Rezeptur Sollwerte - BOOL'
   Button "Button_3" at 160,555 size 78x45; TextOff 'Text'; PictureOff "Up_Arrow"
      on Release: function_b9b71300("CPG_Recipe_Management.currentPages[2]", 1)
   Button "Button_4" at 287,555 size 78x45; TextOff 'Text'; PictureOff "Down_Arrow"
      on Release: function_dd21b452("CPG_Recipe_Management.currentPages[2]", 1)
   TextField "Text field_10" at 35,565 size 126x25; Text 'Pg Up/Down / Seite vor/zurück'
   IOField "I/O field_3" at 446,565 size 35x25; FormatPattern 999
      ProcessValue <- "CPG_Recipe_Management.currentPages[2]"
   TextField "Text field_13" at 381,565 size 60x25; Text 'Page # / Seite #'
   TextField "Text field_14" at 488,565 size 32x25; Text 'of / von'
   IOField "I/O field_4" at 534,564 size 37x27; FormatPattern 999
      ProcessValue <- "CPG_Recipe_Management.maxPages[2]"
   TextField "Text field_2" at 35,93 size 115x25; Text 'Setpoint Name / Sollwert-Name'
   TextField "Text field_6" at 243,83 size 72x46; Text 'Current Value Aktueller Wert'
   TextField "Text field_7" at 384,93 size 32x25; Text 'Min'
   TextField "Text field_4" at 506,93 size 36x25; Text 'Max'
   IOField "I/O field_9" at 757,42 size 53x36; FormatPattern 999
      ProcessValue <- "RecipeID_A"
   IOField "I/O field_10" at 883,42 size 53x36; FormatPattern 999
      ProcessValue <- "RecipeID_B"
   IOField "I/O field_11" at 998,42 size 53x36; FormatPattern 999
      ProcessValue <- "RecipeID_C"
   IOField "I/O field_13" at 550,83 size 187x22; FormatPattern ????????????????????
      ProcessValue <- "CurrentRecipeName"
   IOField "I/O field_14" at 907,104 size 187x22; FormatPattern ????????????????????
      ProcessValue <- "RecipeName_C"
   IOField "I/O field_15" at 816,83 size 187x22; FormatPattern ????????????????????
      ProcessValue <- "RecipeName_B"
   IOField "I/O field_16" at 690,103 size 187x23; FormatPattern ????????????????????
      ProcessValue <- "RecipeName_A"
   TextField "Text field_1" at 748,15 size 98x25; Text 'Recipe A / Datensatz A'
   TextField "Text field_3" at 874,15 size 97x25; Text 'Recipe B / Datensatz B'
   TextField "Text field_8" at 989,15 size 97x25; Text 'Recipe C / Datensatz C'
   Group "Group" at 588,37 size 110x46
   TextField "Text field_5" at 588,37 size 88x46; Text 'Current Recipe: Aktueller Datensatz:'
   IOField "I/O field_12" at 663,48 size 35x25; FormatPattern 999
      ProcessValue <- "CurrentRecipeID"

